
                   #IOuMouldEditor_HMI.arShotSet[#IOuMouldEditor_HMI.sSelected.sPS.iPS].Flow[#TiLoop] := #IOuMouldEditor_HMI.sSelected.sPS.arFlow[#TiLoop];
                   //Sum new Flow
                   #OUTrSumFlow := 0;

                   FOR #TiLoop_Flow := 1 TO #TiComponentAmount DO
                       #OUTrSumFlow := #OUTrSumFlow + #IOuMouldEditor_HMI.arShotSet[#IOuMouldEditor_HMI.sSelected.sPS.iPS].Flow[#TiLoop_Flow];
                   END_FOR;

                   // changed flow is not ref comp
                   IF #TiLoop <> #IOuMouldEditor_HMI.sSelected.sPS.RefComponent THEN
                       // New ratio for changed flow
                       #IOuMouldEditor_HMI.sSelected.sPS.arRatio[#TiLoop] := #IOuMouldEditor_HMI.sSelected.sPS.arFlow[#TiLoop] /
                       #IOuMouldEditor_HMI.arShotSet[#IOuMouldEditor_HMI.sSelected.sPS.iPS].Flow[#IOuMouldEditor_HMI.sSelected.sPS.RefComponent] / 100.0;
                       // changed flow is ref comp    
                   ELSE
                       // New ratio for all other flowrates
                       FOR #TiLoop_Flow := 1 TO #TiComponentAmount DO
                           IF #TiLoop_Flow <> #IOuMouldEditor_HMI.sSelected.sPS.RefComponent THEN
                               IF #IOuMouldEditor_HMI.arShotSet[#IOuMouldEditor_HMI.sSelected.sPS.iPS].Flow[#IOuMouldEditor_HMI.sSelected.sPS.RefComponent] <> 0 THEN
                                   #IOuMouldEditor_HMI.sSelected.sPS.arRatio[#TiLoop_Flow] := #IOuMouldEditor_HMI.sSelected.sPS.arFlow[#TiLoop_Flow] /
                                   #IOuMouldEditor_HMI.arShotSet[#IOuMouldEditor_HMI.sSelected.sPS.iPS].Flow[#IOuMouldEditor_HMI.sSelected.sPS.RefComponent] / 100.0;
                               ELSE
                                   #IOuMouldEditor_HMI.sSelected.sPS.arRatio[#TiLoop_Flow] := 0;
                                   #IOuMouldEditor_HMI.sSelected.sPS.arFlow[#TiLoop_Flow] := 0;
                                   #IOuMouldEditor_HMI.arShotSet[#IOuMouldEditor_HMI.sSelected.sPS.iPS].Flow[#TiLoop_Flow] := 0;
                               END_IF;
                           END_IF;
                       END_FOR;
                   END_IF;

                   //Sum new Flow
                   #OUTrSumFlow := 0;

                   FOR #TiLoop_Flow := 1 TO #TiComponentAmount DO
                       #OUTrSumFlow := #OUTrSumFlow + #IOuMouldEditor_HMI.arShotSet[#IOuMouldEditor_HMI.sSelected.sPS.iPS].Flow[#TiLoop_Flow];
                   END_FOR;
                   #IOuMouldEditor_HMI.sCalculatedValues.arTotalFlow[#IOuMouldEditor_HMI.sSelected.sPS.iPS] := #OUTrSumFlow;


                   // Calculate new ratio
                   // SumRatio
                   #OUTrSumRatio := 0;

                   FOR #TiLoop_Ratio := 1 TO #TiComponentAmount DO
                       #OUTrSumRatio := #OUTrSumRatio + #IOuMouldEditor_HMI.sSelected.sPS.arRatio[#TiLoop_Ratio];
                   END_FOR;

                   //  Calculation = 0 -> shot time fixed
                   IF #IOuMouldEditor_HMI.sSelected.iCalculation = 0 THEN
                       #IOuMouldEditor_HMI.arShotSet[#IOuMouldEditor_HMI.sSelected.sPS.iPS].PartWeight := #IOuMouldEditor_HMI.sCalculatedValues.arTotalFlow[#IOuMouldEditor_HMI.sSelected.sPS.iPS] * #IOuMouldEditor_HMI.arShotSet[#IOuMouldEditor_HMI.sSelected.sPS.iPS].FoamingTime;
                   END_IF;
                   // ----

                   //  Calculation = 2 -> weight fixed
                   IF #IOuMouldEditor_HMI.sSelected.iCalculation = 2 THEN
                       IF #IOuMouldEditor_HMI.sCalculatedValues.arTotalFlow[#IOuMouldEditor_HMI.sSelected.sPS.iPS] >= 0 THEN
                           #IOuMouldEditor_HMI.arShotSet[#IOuMouldEditor_HMI.sSelected.sPS.iPS].FoamingTime := #IOuMouldEditor_HMI.arShotSet[#IOuMouldEditor_HMI.sSelected.sPS.iPS].PartWeight / #IOuMouldEditor_HMI.sCalculatedValues.arTotalFlow[#IOuMouldEditor_HMI.sSelected.sPS.iPS];
                       END_IF;
                   END_IF;

                   //  Value changed + Save data for the last cycle to recognize changes of the values
                   #IOuMouldEditor_HMI.sStatusBits.xValueChanged := TRUE;
                   #SuMouldEditor_HMI := #IOuMouldEditor_HMI;
                   EXIT;
                   // ----

               END_IF
               ;
           END_FOR;
       END_REGION
       //_________________________________________________________________________________    
       REGION Pressure - changed
           FOR #TiLoop := 1 TO #TiComponentAmount DO
               IF #IOuMouldEditor_HMI.sSelected.sPS.arPressure[#TiLoop] <> #SuMouldEditor_HMI.sSelected.sPS.arPressure[#TiLoop] THEN

                   #IOuMouldEditor_HMI.arShotSet[#IOuMouldEditor_HMI.sSelected.sPS.iPS].Pressure[#TiLoop] := #IOuMouldEditor_HMI.sSelected.sPS.arPressure[#TiLoop];

                   //  Value changed + Save data for the last cycle to recognize changes of the values
                   #IOuMouldEditor_HMI.sStatusBits.xValueChanged := TRUE;
                   #SuMouldEditor_HMI := #IOuMouldEditor_HMI;
                   EXIT;
                   // ----

               END_IF
               ;
           END_FOR;
       END_REGION
       //_________________________________________________________________________________    
       REGION Reference component - changed
           IF #IOuMouldEditor_HMI.sSelected.sPS.RefComponent <> #SuMouldEditor_HMI.sSelected.sPS.RefComponent THEN

               #IOuMouldEditor_HMI.arShotSet[#IOuMouldEditor_HMI.sSelected.sPS.iPS].RefComponent := #IOuMouldEditor_HMI.sSelected.sPS.RefComponent;

               IF #IOuMouldEditor_HMI.sSelected.sPS.arFlow[#IOuMouldEditor_HMI.sSelected.sPS.RefComponent] = 0 THEN
                   #IOuMouldEditor_HMI.sSelected.sPS.arRatio[#IOuMouldEditor_HMI.sSelected.sPS.RefComponent] := 100.00;
               END_IF;

               // Calculation of flow in "Mixing ratio - changed"
               //  Value changed + Save data for the last cycle to recognize changes of the values
               #IOuMouldEditor_HMI.sStatusBits.xValueChanged := TRUE;
               //#SuMouldEditor_HMI := #IOuMouldEditor_HMI;

           END_IF;
       END_REGION
       //_________________________________________________________________________________    
       REGION Mixing ratio - changed
           FOR #TiLoop := 1 TO #TiComponentAmount DO
               IF #IOuMouldEditor_HMI.sSelected.sPS.arRatio[#TiLoop] <> #SuMouldEditor_HMI.sSelected.sPS.arRatio[#TiLoop] THEN

                   // only change single flow rates!
                   // SumRatio
                   #OUTrSumRatio := 0;

                   FOR #TiLoop_Ratio := 1 TO #TiComponentAmount DO
                       #OUTrSumRatio := #OUTrSumRatio + #IOuMouldEditor_HMI.sSelected.sPS.arRatio[#TiLoop_Ratio];
                   END_FOR;

                   FOR #TiLoop_Flow := 1 TO #TiComponentAmount DO

                       #IOuMouldEditor_HMI.sSelected.sPS.arFlow[#TiLoop_Flow] := #IOuMouldEditor_HMI.sCalculatedValues.arTotalFlow[#IOuMouldEditor_HMI.sSelected.sPS.iPS] /
                       #OUTrSumRatio * #IOuMouldEditor_HMI.sSelected.sPS.arRatio[#TiLoop_Flow];
                       #IOuMouldEditor_HMI.arShotSet[#IOuMouldEditor_HMI.sSelected.sPS.iPS].Flow[#TiLoop_Flow] := #IOuMouldEditor_HMI.sSelected.sPS.arFlow[#TiLoop_Flow];
                   END_FOR;

                   //  Value changed + Save data for the last cycle to recognize changes of the values
                   #IOuMouldEditor_HMI.sStatusBits.xValueChanged := TRUE;
                   #SuMouldEditor_HMI := #IOuMouldEditor_HMI;
                   EXIT;
                   // ----

               END_IF
               ;
           END_FOR;
       END_REGION
       //_________________________________________________________________________________    
       REGION Mixing head - changed
           FOR #TiLoop_PS := 1 TO #TiPartShotAmount DO
               IF #IOuMouldEditor_HMI.arShotSet[#TiLoop_PS].MHNo <> #SuMouldEditor_HMI.arShotSet[#TiLoop_PS].MHNo THEN
                   // Check if ref comp is available at this MH. Reset all values for not used components            

                   IF #RefComp > #TiComponentAmount THEN
                       #IOuMouldEditor_HMI.arShotSet[#TiLoop_PS].RefComponent := 1;
                   END_IF;

                   IF #TiComponentAmount < 6 THEN
                       FOR #TiLoop := #TiComponentAmount + 1 TO 6 DO
                           #IOuMouldEditor_HMI.arShotSet[#TiLoop_PS].Pressure[#TiLoop] := 0;
                           #IOuMouldEditor_HMI.arShotSet[#TiLoop_PS].Flow[#TiLoop] := 0;
                       END_FOR;
                   END_IF;
                   //  Value changed + Save data for the last cycle to recognize changes of the values
                   #IOuMouldEditor_HMI.sStatusBits.xValueChanged := TRUE;
                   #SuMouldEditor_HMI := #IOuMouldEditor_HMI;
                   EXIT;
                   // ----

               END_IF;
           END_FOR;
       END_REGION
       //_________________________________________________________________________________    
       REGION Two point adjust changed
           // IF #IOuMouldEditor_HMI.sSelected.sPS."2PoinMovement_Comp01" <> #SuMouldEditor_HMI.sSelected.sPS."2PoinMovement_Comp01" OR
           //     #IOuMouldEditor_HMI.sSelected.sPS."2PoinMovement_Comp02" <> #SuMouldEditor_HMI.sSelected.sPS."2PoinMovement_Comp02" OR
           //     #IOuMouldEditor_HMI.sSelected.sPS."2PoinMovement_Comp03" <> #SuMouldEditor_HMI.sSelected.sPS."2PoinMovement_Comp03" OR
           //     #IOuMouldEditor_HMI.sSelected.sPS."2PoinMovement_Comp04" <> #SuMouldEditor_HMI.sSelected.sPS."2PoinMovement_Comp04" OR
           //     #IOuMouldEditor_HMI.sSelected.sPS."2PoinMovement_Comp05" <> #SuMouldEditor_HMI.sSelected.sPS."2PoinMovement_Comp05" OR
           //     #IOuMouldEditor_HMI.sSelected.sPS."2PoinMovement_Comp06" <> #SuMouldEditor_HMI.sSelected.sPS."2PoinMovement_Comp06"
           // THEN
           //     #IOuMouldEditor_HMI.arShotSet[#IOuMouldEditor_HMI.sSelected.sPS.iPS]."2PoinMovement_Comp01" := #IOuMouldEditor_HMI.sSelected.sPS."2PoinMovement_Comp01";
           //     #IOuMouldEditor_HMI.arShotSet[#IOuMouldEditor_HMI.sSelected.sPS.iPS]."2PoinMovement_Comp02" := #IOuMouldEditor_HMI.sSelected.sPS."2PoinMovement_Comp02";
           //     #IOuMouldEditor_HMI.arShotSet[#IOuMouldEditor_HMI.sSelected.sPS.iPS]."2PoinMovement_Comp03" := #IOuMouldEditor_HMI.sSelected.sPS."2PoinMovement_Comp03";
           //     #IOuMouldEditor_HMI.arShotSet[#IOuMouldEditor_HMI.sSelected.sPS.iPS]."2PoinMovement_Comp04" := #IOuMouldEditor_HMI.sSelected.sPS."2PoinMovement_Comp04";
           //     #IOuMouldEditor_HMI.arShotSet[#IOuMouldEditor_HMI.sSelected.sPS.iPS]."2PoinMovement_Comp05" := #IOuMouldEditor_HMI.sSelected.sPS."2PoinMovement_Comp05";
           //     #IOuMouldEditor_HMI.arShotSet[#IOuMouldEditor_HMI.sSelected.sPS.iPS]."2PoinMovement_Comp06" := #IOuMouldEditor_HMI.sSelected.sPS."2PoinMovement_Comp06";

           //     //  Value changed + Save data for the last cycle to recognize changes of the values
           //     #IOuMouldEditor_HMI.sStatusBits.xValueChanged := TRUE;
           //     #SuMouldEditor_HMI := #IOuMouldEditor_HMI;
           //     // ----
           // END_IF;
       END_REGION
       //_________________________________________________________________________________    
       REGION Values in shot settings - changed
           FOR #TiLoop_PS := 1 TO #TiPartShotAmount DO
               IF #IOuMouldEditor_HMI.arShotSet[#TiLoop_PS].MHNo <> #SuMouldEditor_HMI.arShotSet[#TiLoop_PS].MHNo OR
                   #IOuMouldEditor_HMI.arShotSet[#TiLoop_PS].CP_ThrottleGap <> #SuMouldEditor_HMI.arShotSet[#TiLoop_PS].CP_ThrottleGap OR
                   #IOuMouldEditor_HMI.arShotSet[#TiLoop_PS].CP_ThrottleGap <> #SuMouldEditor_HMI.arShotSet[#TiLoop_PS].CP_ThrottleGap OR
                   #IOuMouldEditor_HMI.arShotSet[#TiLoop_PS].PartShotDisable <> #SuMouldEditor_HMI.arShotSet[#TiLoop_PS].PartShotDisable OR
                   #IOuMouldEditor_HMI.arShotSet[#TiLoop_PS].CPMoveAfterShot <> #SuMouldEditor_HMI.arShotSet[#TiLoop_PS].CPMoveAfterShot OR
                   #IOuMouldEditor_HMI.arShotSet[#TiLoop_PS].PartCounter <> #SuMouldEditor_HMI.arShotSet[#TiLoop_PS].PartCounter
               THEN

                   //  Value changed + Save data for the last cycle to recognize changes of the values
                   #IOuMouldEditor_HMI.sStatusBits.xValueChanged := TRUE;
                   #SuMouldEditor_HMI := #IOuMouldEditor_HMI;
                   EXIT;
                   // ----

               END_IF
               ;
           END_FOR;
       END_REGION
       //_________________________________________________________________________________    
       REGION Partial shot number -> copy all data
           FOR #TiLoop := 1 TO #TiComponentAmount DO
               #IOuMouldEditor_HMI.sSelected.sPS.arFlow[#TiLoop] := #IOuMouldEditor_HMI.arShotSet[#IOuMouldEditor_HMI.sSelected.sPS.iPS].Flow[#TiLoop];
               #IOuMouldEditor_HMI.sSelected.sPS.arPressure[#TiLoop] := #IOuMouldEditor_HMI.arShotSet[#IOuMouldEditor_HMI.sSelected.sPS.iPS].Pressure[#TiLoop];
           END_FOR;
       END_REGION
       //_________________________________________________________________________________    
       REGION Reference component = 100%
           #RefComp := LIMIT(MN := 1, IN := #IOuMouldEditor_HMI.sSelected.sPS.RefComponent, MX := #TiComponentAmount);
           #IOuMouldEditor_HMI.sSelected.sPS.RefComponent := #RefComp;
           #TrFlowRefComp := #IOuMouldEditor_HMI.sSelected.sPS.arFlow[#IOuMouldEditor_HMI.sSelected.sPS.RefComponent];
       END_REGION
       //_________________________________________________________________________________    
       REGION Calculate ration out OF flow rate
           FOR #TiLoop := 1 TO #TiComponentAmount DO
               IF #TiLoop = #IOuMouldEditor_HMI.sSelected.sPS.RefComponent THEN
                   #IOuMouldEditor_HMI.sSelected.sPS.arRatio[#TiLoop] := 100.00;
               ELSE
                   IF #TrFlowRefComp > 00 THEN
                       #IOuMouldEditor_HMI.sSelected.sPS.arRatio[#TiLoop] := #IOuMouldEditor_HMI.sSelected.sPS.arFlow[#TiLoop] /
                       #TrFlowRefComp * 100.0;
                   END_IF;
               END_IF;
           END_FOR;
       END_REGION
       //_________________________________________________________________________________    
       #IOuMouldEditor_HMI.sSelected.sPS.RefComponent := #IOuMouldEditor_HMI.arShotSet[#IOuMouldEditor_HMI.sSelected.sPS.iPS].RefComponent;
       //_________________________________________________________________________________    
       REGION Safe changes
           // Check min/max shot time and max flowrates for each component. If out of range ask for change or discard changes   
           IF #IOuMouldEditor_HMI.sStatusBits.xSafeChanges THEN
               FOR #TiLoop_PS := 1 TO #TiPartShotAmount DO
                   // check total flow or total weight is zero
                   IF #IOuMouldEditor_HMI.sCalculatedValues.arTotalFlow[#TiLoop_PS] = 0 OR #IOuMouldEditor_HMI.arShotSet[#TiLoop_PS].PartWeight = 0 THEN
                       #IOuMouldEditor_HMI.sStatusBits.xFaultValuesnotvalid := TRUE;
                   END_IF;
                   // check foaming time for all partshots
                   IF #IOuMouldEditor_HMI.arShotSet[#TiLoop_PS].FoamingTime < "InterfaceVisu".MinShottime OR #IOuMouldEditor_HMI.arShotSet[#TiLoop_PS].FoamingTime > "InterfaceVisu".MaxShottime THEN
                       #IOuMouldEditor_HMI.sStatusBits.xFaultValuesnotvalid := TRUE;
                   END_IF;
                   // check flow rate for all part shots
                   FOR #TiLoop_Flow := 1 TO #TiComponentAmount DO
                       // Maximum flow rate limit reached
                       IF #IOuMouldEditor_HMI.arShotSet[#TiLoop_PS].Flow[#TiLoop_Flow] > "InterfaceVisu".MaxFlow[#TiLoop_Flow] THEN
                           #IOuMouldEditor_HMI.sStatusBits.xFaultValuesnotvalid := TRUE;
                       END_IF;
                       // Minimum flow rate limit reached
                       IF #IOuMouldEditor_HMI.arShotSet[#TiLoop_PS].Flow[#TiLoop_Flow] < "InterfaceVisu".MinFlow[#TiLoop_Flow] AND
                           #IOuMouldEditor_HMI.arShotSet[#TiLoop_PS].Flow[#TiLoop_Flow] <> 0 THEN
                           #IOuMouldEditor_HMI.sStatusBits.xFaultValuesnotvalid := TRUE;
                       END_IF;

                   END_FOR;

               END_FOR;
               #IOuMouldEditor_HMI.sStatusBits.xSafeChanges := FALSE;

               IF #IOuMouldEditor_HMI.sStatusBits.xFaultValuesnotvalid = FALSE THEN
                   #IOuMouldEditor_HMI.sStatusBits.xValueChanged := FALSE;
                   #IOuMouldEditor_HMI.sStatusBits.xSafeChanges := FALSE;
                   #IOuMouldEditor_HMI.sStatusBits.xDiscardChanges := FALSE;

                   FOR #TiLoop_PS := 1 TO #TiPartShotAmount DO
                       // When the selected Tool less or equal 100 is, transfer the values to DB925
                       IF #IOuMouldEditor_HMI.sSelected.iTool <= "AmountToolsDB" THEN
                           "DB925_ShotData_1".Tool[#IOuMouldEditor_HMI.sSelected.iTool].Shot[#TiLoop_PS] := #IOuMouldEditor_HMI.arShotSet[#TiLoop_PS];
                       END_IF;
                       // When the selected Tool bigger than 100 and less or equal 200 is, transfer the values to DB926
                       IF #IOuMouldEditor_HMI.sSelected.iTool > "AmountToolsDB" AND #IOuMouldEditor_HMI.sSelected.iTool <= (2*"AmountToolsDB") THEN
                           "DB926_ShotData_2".Tool[#IOuMouldEditor_HMI.sSelected.iTool-"AmountToolsDB"].Shot[#TiLoop_PS] := #IOuMouldEditor_HMI.arShotSet[#TiLoop_PS];
                       END_IF;
                   END_FOR;

                   "DB930_Tools".Tool[#IOuMouldEditor_HMI.sSelected.iTool] := #IOuMouldEditor_HMI.uTools;
               END_IF;
           END_IF;
       END_REGION
       //_________________________________________________________________________________    
       REGION Delete program
           IF #IOuMouldEditor_HMI.sStatusBits.xDeleteProgram THEN
               #IOuMouldEditor_HMI.sStatusBits.xDeleteProgram := false;
               "FC4_Check_allocation"(Selected_tool:=#IOuMouldEditor_HMI.sSelected.iTool,
                                      Delete_not_allowed=>#IOuMouldEditor_HMI.sStatusBits.xFaultDeleteProgram);

               IF NOT #IOuMouldEditor_HMI.sStatusBits.xFaultDeleteProgram THEN
                   #IOuMouldEditor_HMI.uTools.PartShot_Amount := 0;
                   #Nullbyte := 0;
                   // Delete tool data
                   // When the selected Tool less or equal 100 is, transfer the values to DB925
                   IF #IOuMouldEditor_HMI.sSelected.iTool <= "AmountToolsDB" THEN
                       #Retval := FILL(BVAL := #Nullbyte, BLK => "DB925_ShotData_1".Tool[#IOuMouldEditor_HMI.sSelected.iTool]);
                   END_IF;
                   // When the selected Tool bigger than 100 and less or equal 200 is, transfer the values to DB926
                   IF #IOuMouldEditor_HMI.sSelected.iTool > "AmountToolsDB" AND #IOuMouldEditor_HMI.sSelected.iTool <= (2 * "AmountToolsDB") THEN
                       #Retval := FILL(BVAL := #Nullbyte, BLK => "DB926_ShotData_2".Tool[#IOuMouldEditor_HMI.sSelected.iTool-"AmountToolsDB"]);
                   END_IF;

                   #Retval := FILL(BVAL := #Nullbyte, BLK => "DB930_Tools".Tool[#IOuMouldEditor_HMI.sSelected.iTool]);
                   #Retval := FILL(BVAL := #Nullbyte, BLK => #IOuMouldEditor_HMI.arShotSet);
                   "DB930_Tools".Tool[#IOuMouldEditor_HMI.sSelected.iTool].tool_name := '';
               END_IF;

           END_IF;
       END_REGION
       //_________________________________________________________________________________    
       REGION Save data FOR the last cycle TO recognize changes OF the values
           #SuMouldEditor_HMI := #IOuMouldEditor_HMI;
       END_REGION
       //_________________________________________________________________________________    
       REGION Visibility OF part shots AND "grey" fields FOR NOT changing settings
           // Column
           // Column - shot time blocked
           IF #IOuMouldEditor_HMI.sSelected.iCalculation = 0 THEN   // Statement section REGION
               #IOuMouldEditor_HMI.sColumn.iShotTime := #IOuMouldEditor_HMI.uTools.PartShot_Amount;
           ELSE
               #IOuMouldEditor_HMI.sColumn.iShotTime := 0;
           END_IF;

           // Column - total flow blocked
           IF #IOuMouldEditor_HMI.sSelected.iCalculation = 1 THEN   // Statement section REGION
               #IOuMouldEditor_HMI.sColumn.iTotalFlow := #IOuMouldEditor_HMI.uTools.PartShot_Amount;
           ELSE
               #IOuMouldEditor_HMI.sColumn.iTotalFlow := 0;
           END_IF;

           // Column - total weight blocked
           IF #IOuMouldEditor_HMI.sSelected.iCalculation = 2 THEN   // Statement section REGION
               #IOuMouldEditor_HMI.sColumn.iTotalWeight := #IOuMouldEditor_HMI.uTools.PartShot_Amount;
           ELSE
               #IOuMouldEditor_HMI.sColumn.iTotalWeight := 0;
           END_IF;

           // Row - Visibility of change partial shot
           FOR #TiLoop := 1 TO "AmountPartShots" DO
               IF #TiLoop <> #IOuMouldEditor_HMI.sSelected.sPS.iPS AND
                   #TiLoop <= BYTE_TO_INT(#IOuMouldEditor_HMI.uTools.PartShot_Amount)
               THEN
                   #IOuMouldEditor_HMI.sRow.arChangePartialShot[#TiLoop] := TRUE;
               ELSE
                   #IOuMouldEditor_HMI.sRow.arChangePartialShot[#TiLoop] := FALSE;
               END_IF;

           END_FOR;
       END_REGION
   END_IF;
END_FUNCTION_BLOCK

FUNCTION_BLOCK "FB009_Faults"   // FB9, STL
TITLE = Faults indication of machines and plant
{ S7_Optimized_Access := 'FALSE' }
AUTHOR : KT242
VERSION : 0.1
   VAR_TEMP
      Stoe_Quitt : Bool;
      Quitt : Bool;
   END_VAR
BEGIN

REGION Network 1
   //      O     "E0.4QuitFault"
   //      O     "Tag_7"
   //      =     "E0.4QuitFault"
END_REGION

REGION Network 2: Bits of fault levels
         A     "DB009_Faults".Faults_FKT_Grp_1_M1;
         =     "DB009_Faults".Fault_State_Grp_1_M1;
         A     "DB009_Faults".Faults_FKT_Grp_2_M1;
         =     "DB009_Faults".Fault_State_Grp_2_M1;
         A     "DB009_Faults".Faults_FKT_Grp_3_M1;
         =     "DB009_Faults".Fault_State_Grp_3_M1;

         A     "DB009_Faults".Faults_FKT_Grp_1_M2;
         =     "DB009_Faults".Fault_State_Grp_1_M2;
         A     "DB009_Faults".Faults_FKT_Grp_2_M2;
         =     "DB009_Faults".Fault_State_Grp_2_M2;
         A     "DB009_Faults".Faults_FKT_Grp_3_M2;
         =     "DB009_Faults".Fault_State_Grp_3_M2;

         CLR;
         =     "DB009_Faults".Fault_State_Grp_1_M3;
         =     "DB009_Faults".Fault_State_Grp_2_M3;
         =     "DB009_Faults".Fault_State_Grp_3_M3;
         =     "DB009_Faults".Fault_State_Grp_1_M4;
         =     "DB009_Faults".Fault_State_Grp_2_M4;
         =     "DB009_Faults".Fault_State_Grp_3_M4;

         A     "DB009_Faults".Faults_FKT_Grp_1_ExtP;
         =     "DB009_Faults".Fault_State_Grp_1_ExtP;
         A     "DB009_Faults".Faults_FKT_Grp_2_ExtP;
         =     "DB009_Faults".Fault_State_Grp_2_ExtP;
         A     "DB009_Faults".Faults_FKT_Grp_3_ExtP;
         =     "DB009_Faults".Fault_State_Grp_2_ExtP;

         O     "T_QuitFault";
         O     "FRA_KM_Quitt";
         =     #Quitt;

         CALL  "FC089_quit_Faults"
         ( IN_Button_Acknowledge    := #Quitt,  //"T_QuitFault"
           IN_Button_Horn_Off       := FALSE,  // "E0.4QuitFault"
           IN_First_PLC_cycle       := "Flag_Erster_SPS_Zyklus",
           IN_IndicatorLampTest     := "DB619_State_MPart".Operationmode[1].Lamptest,
           IN_Fault_Grp_1_active_M1 := "DB009_Faults".Fault_State_Grp_1_M1,
           IN_Fault_Grp_2_active_M1 := "DB009_Faults".Fault_State_Grp_2_M1,
           IN_Fault_Grp_3_active_M1 := "DB009_Faults".Fault_State_Grp_3_M1,
           IN_Fault_Grp_1_active_M2 := "DB009_Faults".Fault_State_Grp_1_M2,
           IN_Fault_Grp_2_active_M2 := "DB009_Faults".Fault_State_Grp_2_M2,
           IN_Fault_Grp_3_active_M2 := "DB009_Faults".Fault_State_Grp_3_M2,
           IN_Fault_Grp_1_active_M3 := "DB009_Faults".Fault_State_Grp_1_M3,
           IN_Fault_Grp_2_active_M3 := "DB009_Faults".Fault_State_Grp_2_M3,
           IN_Fault_Grp_3_active_M3 := "DB009_Faults".Fault_State_Grp_3_M3,
           IN_Fault_Grp_1_active_M4 := "DB009_Faults".Fault_State_Grp_1_M4,
           IN_Fault_Grp_2_active_M4 := "DB009_Faults".Fault_State_Grp_2_M4,
           IN_Fault_Grp_3_active_M4 := "DB009_Faults".Fault_State_Grp_3_M4,
           IN_Fault_Grp_1_active_AP := "DB009_Faults".Fault_State_Grp_1_ExtP,
           IN_Fault_Grp_2_active_AP := "DB009_Faults".Fault_State_Grp_2_ExtP,
           IN_Fault_Grp_3_active_AP := "DB009_Faults".Fault_State_Grp_3_ExtP,
           OUT_acoustical_indicator := "H_Fault_horn_M1",
           OUT_optical_indicator    := "H_Fault_lamp_M1",
           IO_Fault_changed_M1      := "DB009_Faults".Faultschanging_M1,
           IO_Fault_changed_M2      := "DB009_Faults".Faultschanging_M2,
           IO_Fault_changed_M3      := "DB009_Faults".Faultschanging_M3,
           IO_Fault_changed_M4      := "DB009_Faults".Faultschanging_M4,
           IO_Fault_changed_AP      := "DB009_Faults".Faultschanging_ExtP,
           IO_Horn                  := "DB009_Faults".HF_Horn,
           IO_Reset_fault_Grp       := "DB009_Faults".Faults_Reset_Group,
           IO_Reset_fault_Fkt       := "DB009_Faults".Faults_Reset_FKT_M1,
           IO_Quit_Edge             := "DB009_Faults".HF_Faults_Quit
         );
   //-----
         O     "DB009_Faults".Fault_State_Grp_1_M1;
         O     "DB009_Faults".Fault_State_Grp_2_M1;
         O     "DB009_Faults".Fault_State_Grp_3_M1;
         O     "DB009_Faults".Fault_State_Grp_1_M2;
         O     "DB009_Faults".Fault_State_Grp_2_M2;
         O     "DB009_Faults".Fault_State_Grp_3_M2;
         O     "DB009_Faults".Fault_State_Grp_1_M3;
         O     "DB009_Faults".Fault_State_Grp_2_M3;
         O     "DB009_Faults".Fault_State_Grp_3_M3;
         O     "DB009_Faults".Fault_State_Grp_1_M4;
         O     "DB009_Faults".Fault_State_Grp_2_M4;
         O     "DB009_Faults".Fault_State_Grp_3_M4;
         O     "DB009_Faults".Fault_State_Grp_1_ExtP;
         O     "DB009_Faults".Fault_State_Grp_2_ExtP;
         O     "DB009_Faults".Fault_State_Grp_2_ExtP;
         =     "DB009_Faults".Fault_State_Grp_1_3_Exist;
   //-----
         A     "DB009_Faults".Faults_Reset_FKT_M1;
         S     "DB009_Faults".HF_FaultsQuitOB35;
   //-----
         A     "DB009_Faults".Faults_Reset_Group;
         R     "DB009_Faults".Faults_FKT_Grp_1_M1;
         R     "DB009_Faults".Faults_FKT_Grp_2_M1;
         R     "DB009_Faults".Faults_FKT_Grp_3_M1;
         R     "DB009_Faults".Faults_FKT_Grp_1_M2;
         R     "DB009_Faults".Faults_FKT_Grp_2_M2;
         R     "DB009_Faults".Faults_FKT_Grp_3_M2;
         R     "DB009_Faults".Faults_FKT_Grp_1_M3;
         R     "DB009_Faults".Faults_FKT_Grp_2_M3;
         R     "DB009_Faults".Faults_FKT_Grp_3_M3;
         R     "DB009_Faults".Faults_FKT_Grp_1_M4;
         R     "DB009_Faults".Faults_FKT_Grp_2_M4;
         R     "DB009_Faults".Faults_FKT_Grp_3_M4;
         R     "DB009_Faults".Faults_FKT_Grp_1_ExtP;
         R     "DB009_Faults".Faults_FKT_Grp_2_ExtP;
         R     "DB009_Faults".Faults_FKT_Grp_3_ExtP;
   //-----
END_REGION

REGION Network 3: General faults of machines
         CALL  "FC081_FaultsGen"
         ( IN_Erster_SPS_Zyklus := "Flag_Erster_SPS_Zyklus"
         );
END_REGION

REGION Network 4: Faults Profibus
         CALL  "FC082_FaultProfiBus";
END_REGION

REGION Network 5: Lamp machine ok for foaming
         O     "H_Ready_for_Operation_M1";
         O     "H_Ready_for_Operation_M2";
         =     "H_Ready_for_Operation";
END_REGION

REGION Network 6: Signalshow fault massages and messages at visu
         O     "DB009_Faults".NewMessage_M1;
         O     "DB009_Faults".GoneMessage_M1;
         O     "DB009_Faults".Faultschanging_M1;
         O     "DB009_Faults".Faults_Reset_FKT_M1;
         AN    "DB009_Faults".MessageChangedToVisu;
         S     "DB009_Faults".MessageChangedToVisu;
         R     "DB009_Faults".NewMessage_M1;
         R     "DB009_Faults".GoneMessage_M1;
         R     "DB009_Faults".MessageChangedNext;

         O     "DB009_Faults".NewMessage_M1;
         O     "DB009_Faults".GoneMessage_M1;
         O     "DB009_Faults".Faultschanging_M1;
         O     "DB009_Faults".Faults_Reset_FKT_M1;
         A     "DB009_Faults".MessageChangedToVisu;
         S     "DB009_Faults".MessageChangedNext;
END_REGION
END_FUNCTION_BLOCK

FUNCTION_BLOCK "FB011_OP_CirceMode_M1"   // FB11, STL
TITLE = Operation mode and cycle mode of machine 01
{ S7_Optimized_Access := 'FALSE' }
AUTHOR : KT242
VERSION : 0.1
   VAR_TEMP
      Temp_Release_HP : Bool;
      Temp_ShotPreperation : Bool;
      Temp_Automatic_MH1 : Bool;
      Temp_HPCirc_aft_shot_MH1 : Bool;
      Temp_HF_LP_circ : Bool;
      Temp_TestMode : Bool;
      Temp_TestA : Bool;
      Temp_TestB : Bool;
      Temp_H_TestA : Bool;
      Temp_H_TestB : Bool;
      Dummy : Bool;
   END_VAR
BEGIN

REGION Network 1: State switch service/ operation
         L     0;
         T     "DB614_MH_State".MH_Status[1].State_Service;
         T     "DB614_MH_State".MH_Status[2].State_Service;
         T     "DB614_MH_State".MH_Status[3].State_Service;
         T     "DB614_MH_State".MH_Status[4].State_Service;
         T     "DB614_MH_State".MH_Status[5].State_Service;
         T     "DB614_MH_State".MH_Status[6].State_Service;
         T     "DB614_MH_State".MH_Status[7].State_Service;
         T     "DB614_MH_State".MH_Status[8].State_Service;
         T     "DB614_MH_State".MH_Status[8].State_Service;
         T     "DB614_MH_State".MH_Status[9].State_Service;
         T     "DB614_MH_State".MH_Status[10].State_Service;
         T     "DB614_MH_State".MH_Status[11].State_Service;
         T     "DB614_MH_State".MH_Status[12].State_Service;
   //-----
         A     "DB614_MH_State".MH_Status[1].Switch_Service_ON_OFF;
         JCN   NoServ_MH01;
         L     1;
         T     "DB614_MH_State".MH_Status[1].State_Service;
   NoServ_MH01:NOP   0;
   //-----
         A     "DB614_MH_State".MH_Status[2].Switch_Service_ON_OFF;
         JCN   NoServ_MH02;
         L     1;
         T     "DB614_MH_State".MH_Status[2].State_Service;
   NoServ_MH02:NOP   0;
   //-----
         A     "DB614_MH_State".MH_Status[3].Switch_Service_ON_OFF;
         JCN   NoServ_MH03;
         L     1;
         T     "DB614_MH_State".MH_Status[3].State_Service;
   NoServ_MH03:NOP   0;
   //-----
         A     "DB614_MH_State".MH_Status[4].Switch_Service_ON_OFF;
         JCN   NoServ_MH04;
         L     1;
         T     "DB614_MH_State".MH_Status[4].State_Service;
   NoServ_MH04:NOP   0;
   //-----
         A     "DB614_MH_State".MH_Status[5].Switch_Service_ON_OFF;
         JCN   NoServ_MH05;
         L     1;
         T     "DB614_MH_State".MH_Status[5].State_Service;
   NoServ_MH05:NOP   0;
   //-----
         A     "DB614_MH_State".MH_Status[6].Switch_Service_ON_OFF;
         JCN   NoServ_MH06;
         L     1;
         T     "DB614_MH_State".MH_Status[6].State_Service;
   NoServ_MH06:NOP   0;
   //-----
         A     "DB614_MH_State".MH_Status[7].Switch_Service_ON_OFF;
         JCN   NoServ_MH07;
         L     1;
         T     "DB614_MH_State".MH_Status[7].State_Service;
   NoServ_MH07:NOP   0;
   //-----
         A     "DB614_MH_State".MH_Status[8].Switch_Service_ON_OFF;
         JCN   NoServ_MH08;
         L     1;
         T     "DB614_MH_State".MH_Status[8].State_Service;
   NoServ_MH08:NOP   0;
   //-----
         A     "DB614_MH_State".MH_Status[9].Switch_Service_ON_OFF;
         JCN   NoServ_MH09;
         L     1;
         T     "DB614_MH_State".MH_Status[9].State_Service;
   NoServ_MH09:NOP   0;
   //-----
         A     "DB614_MH_State".MH_Status[10].Switch_Service_ON_OFF;
         JCN   NoServ_MH10;
         L     1;
         T     "DB614_MH_State".MH_Status[10].State_Service;
   NoServ_MH10:NOP   0;
   //-----
         A     "DB614_MH_State".MH_Status[11].Switch_Service_ON_OFF;
         JCN   NoServ_MH11;
         L     1;
         T     "DB614_MH_State".MH_Status[11].State_Service;
   NoServ_MH11:NOP   0;
   //-----
         A     "DB614_MH_State".MH_Status[12].Switch_Service_ON_OFF;
         JCN   NoServ_MH12;
         L     1;
         T     "DB614_MH_State".MH_Status[12].State_Service;
   NoServ_MH12:NOP   0;
   //-----
END_REGION

REGION Network 2: Switch operation mode ->ON -> with foam to open mixinghead (extarnel)

         A     "DB619_State_MPart".SWU[1].Open_SWU."01";
         A     "DB614_MH_State".MH_Status[1].Switch_Service_ON_OFF;
         O;
         A     "DB619_State_MPart".SWU[1].Open_SWU."02";
         A     "DB614_MH_State".MH_Status[2].Switch_Service_ON_OFF;
         O;
         A     "DB619_State_MPart".SWU[1].Open_SWU."03";
         A     "DB614_MH_State".MH_Status[3].Switch_Service_ON_OFF;
         O;
         A     "DB619_State_MPart".SWU[1].Open_SWU."04";
         A     "DB614_MH_State".MH_Status[4].Switch_Service_ON_OFF;
         O;
         A     "DB619_State_MPart".SWU[1].Open_SWU."05";
         A     "DB614_MH_State".MH_Status[5].Switch_Service_ON_OFF;
         O;
         A     "DB619_State_MPart".SWU[1].Open_SWU."06";
         A     "DB614_MH_State".MH_Status[6].Switch_Service_ON_OFF;
         O;
         A     "DB619_State_MPart".SWU[1].Open_SWU."07";
         A     "DB614_MH_State".MH_Status[7].Switch_Service_ON_OFF;
         O;
         A     "DB619_State_MPart".SWU[1].Open_SWU."08";
         A     "DB614_MH_State".MH_Status[8].Switch_Service_ON_OFF;
         O;
         A     "DB619_State_MPart".SWU[1].Open_SWU."09";
         A     "DB614_MH_State".MH_Status[9].Switch_Service_ON_OFF;
         O;
         A     "DB619_State_MPart".SWU[1].Open_SWU."10";
         A     "DB614_MH_State".MH_Status[10].Switch_Service_ON_OFF;
         O;
         A     "DB619_State_MPart".SWU[1].Open_SWU."11";
         A     "DB614_MH_State".MH_Status[11].Switch_Service_ON_OFF;
         O;
         A     "DB619_State_MPart".SWU[1].Open_SWU."12";
         A     "DB614_MH_State".MH_Status[12].Switch_Service_ON_OFF;
         =     "DB619_State_MPart".Operationmode[1].SwitchOperation;
END_REGION

REGION Network 3: Test shot Sonder
         L     0;
         T     "DB614_MH_State".MH_Status[1].State_Testshot_A;
         T     "DB614_MH_State".MH_Status[1].State_Testshot_B;

         AN    "DB123_MH_IO_Signals".MH[1].IN.MH_Manual_Mode;
         R     "DB614_MH_State".MH_Status[1].Switch_Testshot_A_ON_OFF;
         R     "DB614_MH_State".MH_Status[1].Switch_Testshot_B_ON_OFF;

         A     "DB614_MH_State".MH_Status[1].Switch_Testshot_A_ON_OFF;
         JCN   TestA_MH01;
         L     1;
         T     "DB614_MH_State".MH_Status[1].State_Testshot_A;
         L     0;
         T     "DB614_MH_State".MH_Status[1].State_Testshot_B;
   TestA_MH01:NOP   0;

         A     "DB614_MH_State".MH_Status[1].Switch_Testshot_B_ON_OFF;
         JCN   TestB_MH01;
         L     1;
         T     "DB614_MH_State".MH_Status[1].State_Testshot_B;
         L     0;
         T     "DB614_MH_State".MH_Status[1].State_Testshot_A;
   TestB_MH01:NOP   0;

         A     "DB614_MH_State".MH_Status[1].Switch_Testshot_A_ON_OFF;
         O     "DB614_MH_State".MH_Status[1].Switch_Testshot_B_ON_OFF;
         =     #Temp_TestMode;

         A     "DB614_MH_State".MH_Status[1].Switch_Testshot_A_ON_OFF;
         A     "DB123_MH_IO_Signals".MH[1].IN.MH_Start;
         =     #Temp_TestA;

         A     "DB614_MH_State".MH_Status[1].Switch_Testshot_B_ON_OFF;
         A     "DB123_MH_IO_Signals".MH[1].IN.MH_Start;
         =     #Temp_TestB;

         A     "DB009_Faults".Faults_FKT_Grp_1_M1;
         L     s5t#3s;
         SP    "TM_Group1_Fault";

         A     #Temp_TestMode;
         A     "DB619_State_MPart".Cycle[1].running;
         AN    "DB614_MH_State".MH_Status[1].Switch_Testshot_A_ON_OFF;
         O     "DB123_MH_IO_Signals".MH[1].OUT.MH.V_LowPressure_Circ_MH;
         O     "TM_Group1_Fault";
   //      NOT
         =     "V_Bypass_C1";

         A     #Temp_TestMode;
         A     "DB619_State_MPart".Cycle[1].running;
         AN    "DB614_MH_State".MH_Status[1].Switch_Testshot_B_ON_OFF;
         O     "DB123_MH_IO_Signals".MH[1].OUT.MH.V_LowPressure_Circ_MH;
         O     "TM_Group1_Fault";
   //      NOT
         =     "V_Bypass_C2";
END_REGION

REGION Network 4: Auslitern
         CALL  "FC115_Testen"
         ( IN_Betriebsart_Testen   := "DB619_State_MPart".Operationmode[1].Test,
           IN_Betriebsart_Betrieb  := "DB619_State_MPart".Operationmode[1].Operation,
           IN_Lampentest           := FALSE,
           IN_Start_Testen_K1      := #Temp_TestA,
           IN_Start_Testen_K2      := #Temp_TestB,
           IN_Start_Testen_K3      := FALSE,
           IN_Start_Testen_K4      := FALSE,
           IN_Stop_Testen          := "DB123_MH_IO_Signals".MH[1].IN.MH_Stop,
           IN_Stoerung_Gruppe_1    := "DB009_Faults".Faults_FKT_Grp_1_M1,
           IN_Zyklus_Freigabe      := "DB619_State_MPart".Cycle[1].Release,
           IN_Zyklus_laeuft        := "DB619_State_MPart".ToolMa[1].StationActive,
           IN_Zyklus_Schuss_laeuft := "DB619_State_MPart".Cycle[1].ShotRuns,
           IN_Imp_Zyklus_Ende      := "DB619_State_MPart".Cycle[1].Pulse_ToolFinished,
           IN_Zyklus_KLZ2_u_ff     := "DB619_State_MPart".Cycle[1].LastStanbyTimeTool,
           OUT_H_Testen_K1         := #Temp_H_TestA,
           OUT_H_Testen_K2         := #Temp_H_TestB,
           OUT_H_Testen_K3         := #Dummy,
           OUT_H_Testen_K4         := #Dummy,
           OUT_V_Testen_K1         := #Dummy,
           OUT_V_Testen_K2         := #Dummy,
           OUT_V_Testen_K3         := #Dummy,
           OUT_V_Testen_K4         := #Dummy,
           IO_Status               := "DB110_Interf_Program_M1".Test_M01
         );
   //
         A     "DB110_Interf_Program_M1".Test_M01.Test_K2;
         =     "Duese_K1_MH01";

         A     "DB110_Interf_Program_M1".Test_M01.Test_K1;
         =     "Duese_K2_MH01";

         A     #Temp_H_TestA;
         O     #Temp_H_TestB;
         =     "DB110_Interf_Program_M1".Test_M01.Spare_0_7;
END_REGION

REGION Network 5: Detecting operation modes
   //-----
         CALL  "FC011_OperationMode"
         ( IN_ContrVoltage        := "Controlvoltage",
           IN_Connection_OK       := TRUE,
           IN_SS_Manual           := "S_OM_Manual",
           IN_SS_Auto             := "S_OM_Auto",
           IN_SS_Test             := #Temp_TestMode,  //"S_OM_Test"
           IN_LampTest            := FALSE,  // "T_Lampentest"
           IN_Cycle_selected      := "DB619_State_MPart".Recirculation[1].Is_selected,
           IN_SS_CylinderService  := "DB619_State_MPart".CylinderManager[1].Cylinderservice,
           IN_Hydraulic_OK        := "DB619_State_MPart".Machine[1].HydStartUp_finished,
           IN_OperationMode_Timer := "TM_OM_M1",
           IO_Status              := "DB619_State_MPart".Operationmode[1]
         );
   //-----
END_REGION

REGION Network 6: High pressure cycle after automatic shot
   //-----
         A     "DB123_MH_IO_Signals".MH[1].IN.MH_Auto_Mode;
         A     "DB619_State_MPart".SWU[1].Open_SWU_allone."01";
   //     CLR
         =     #Temp_Automatic_MH1;
   //-----
         A     "DB619_State_MPart".Cycle[1].ShotRuns;
         A     #Temp_Automatic_MH1;
         L     "DB700_Machine".Machine[1].HP_time_after_shot;
         SF    "TM_HP_after_shot_M1";
   //-----
         O     "TM_HP_after_shot_M1";
   //      CLR
         =     "DB619_State_MPart".Machine[1].HP_after_shot;
   //-----
         A(;
         O     "DB619_State_MPart".Machine[1].HP_after_shot;
         FP    "DB619_State_MPart".Machine[1].Flag_P_HP_after_shot;
         );
         AN    "DB619_State_MPart".Recirculation[1].HP_is_active;
         O;
         A(;
         A     "DB619_State_MPart".Machine[1].HP_after_shot;
         FN    "DB619_State_MPart".Machine[1].Flag_N_HP_after_shot;
         );
         A     "DB619_State_MPart".Recirculation[1].HP_is_active;
         =     #Temp_HPCirc_aft_shot_MH1;
   //-----
         A     #Temp_Automatic_MH1;
         JC    M001;
         L     S5T#0MS;
         CLR;
         SP    "TM_HP_after_shot_M1";
   M001: NOP   0;
   //-----
END_REGION

REGION Network 7: Release of high pressure cycle
         O     "DB619_State_MPart".Machine[1].HP_after_shot;
         ON    "DB619_State_MPart".Cycle[1].running;
         A     "DB619_State_MPart".Operationmode[1].Active;
         AN    "DB009_Faults".Fault_State_Grp_1_M1;
         =     #Temp_Release_HP;
   //-----
END_REGION

REGION Network 8: Select high pressure cycle by PUC08 or mixinghead panel
   //__________________________________________________________________
   // Select high pressure mixinghead 01:
   // ------------------------------------
         O     #Temp_HPCirc_aft_shot_MH1;
         O     "DB123_MH_IO_Signals".MH[1].IN.MH_HP_Circ_MH;
         O     "DB614_MH_State".MH_Status[1].Switch_HP_ON_OFF;
         =     "DB619_State_MPart".Recirculation[1].Button_HP."01";
   //__________________________________________________________________
   //Select high pressure mixinghead 02:
   //------------------------------------
         O     "DB123_MH_IO_Signals".MH[2].IN.MH_HP_Circ_MH;
         O     "DB614_MH_State".MH_Status[2].Switch_HP_ON_OFF;
         =     "DB619_State_MPart".Recirculation[1].Button_HP."02";
   //__________________________________________________________________
   //Select high pressure mixinghead 03:
   //------------------------------------
         O     "DB123_MH_IO_Signals".MH[3].IN.MH_HP_Circ_MH;
         O     "DB614_MH_State".MH_Status[3].Switch_HP_ON_OFF;
         =     "DB619_State_MPart".Recirculation[1].Button_HP."03";
   //__________________________________________________________________
   //Select high pressure mixinghead 04:
   //------------------------------------
         O     "DB123_MH_IO_Signals".MH[4].IN.MH_HP_Circ_MH;
         O     "DB614_MH_State".MH_Status[4].Switch_HP_ON_OFF;
         =     "DB619_State_MPart".Recirculation[1].Button_HP."04";
   //__________________________________________________________________
   //Select high pressure mixinghead 05:
   //------------------------------------
         O     "DB123_MH_IO_Signals".MH[5].IN.MH_HP_Circ_MH;
         O     "DB614_MH_State".MH_Status[5].Switch_HP_ON_OFF;
         =     "DB619_State_MPart".Recirculation[1].Button_HP."05";
   //__________________________________________________________________
   //Select high pressure mixinghead 06:
   //------------------------------------
         O     "DB123_MH_IO_Signals".MH[6].IN.MH_HP_Circ_MH;
         O     "DB614_MH_State".MH_Status[6].Switch_HP_ON_OFF;
         =     "DB619_State_MPart".Recirculation[1].Button_HP."06";
   //__________________________________________________________________
   //Select high pressure mixinghead 07:
   //------------------------------------
         O     "DB123_MH_IO_Signals".MH[7].IN.MH_HP_Circ_MH;
         O     "DB614_MH_State".MH_Status[7].Switch_HP_ON_OFF;
         =     "DB619_State_MPart".Recirculation[1].Button_HP."07";
   //__________________________________________________________________
   //Select high pressure mixinghead 08:
   //------------------------------------
         O     "DB123_MH_IO_Signals".MH[8].IN.MH_HP_Circ_MH;
         O     "DB614_MH_State".MH_Status[8].Switch_HP_ON_OFF;
         =     "DB619_State_MPart".Recirculation[1].Button_HP."08";
   //__________________________________________________________________
   //Select high pressure mixinghead 09:
   //------------------------------------
         O     "DB123_MH_IO_Signals".MH[9].IN.MH_HP_Circ_MH;
         O     "DB614_MH_State".MH_Status[9].Switch_HP_ON_OFF;
         =     "DB619_State_MPart".Recirculation[1].Button_HP."09";
   //__________________________________________________________________
   //Select high pressure mixinghead 10:
   //------------------------------------
         O     "DB123_MH_IO_Signals".MH[10].IN.MH_HP_Circ_MH;
         O     "DB614_MH_State".MH_Status[10].Switch_HP_ON_OFF;
         =     "DB619_State_MPart".Recirculation[1].Button_HP."10";
   //__________________________________________________________________
   //Select high pressure mixinghead 11:
   //------------------------------------
         O     "DB123_MH_IO_Signals".MH[11].IN.MH_HP_Circ_MH;
         O     "DB614_MH_State".MH_Status[11].Switch_HP_ON_OFF;
         =     "DB619_State_MPart".Recirculation[1].Button_HP."11";
   //__________________________________________________________________
   //Select high pressure mixinghead 12:
   //------------------------------------
         O     "DB123_MH_IO_Signals".MH[12].IN.MH_HP_Circ_MH;
         O     "DB614_MH_State".MH_Status[12].Switch_HP_ON_OFF;
         =     "DB619_State_MPart".Recirculation[1].Button_HP."12";
   //__________________________________________________________________
   //
END_REGION

REGION Network 9: Reset the HP switches at the Panel
         SET;
         R     "DB614_MH_State".MH_Status[0].Switch_HP_ON_OFF;
         R     "DB614_MH_State".MH_Status[1].Switch_HP_ON_OFF;
         R     "DB614_MH_State".MH_Status[2].Switch_HP_ON_OFF;
         R     "DB614_MH_State".MH_Status[3].Switch_HP_ON_OFF;
         R     "DB614_MH_State".MH_Status[4].Switch_HP_ON_OFF;
         R     "DB614_MH_State".MH_Status[5].Switch_HP_ON_OFF;
         R     "DB614_MH_State".MH_Status[6].Switch_HP_ON_OFF;
         R     "DB614_MH_State".MH_Status[7].Switch_HP_ON_OFF;
         R     "DB614_MH_State".MH_Status[8].Switch_HP_ON_OFF;
         R     "DB614_MH_State".MH_Status[9].Switch_HP_ON_OFF;
         R     "DB614_MH_State".MH_Status[10].Switch_HP_ON_OFF;
         R     "DB614_MH_State".MH_Status[11].Switch_HP_ON_OFF;
         R     "DB614_MH_State".MH_Status[12].Switch_HP_ON_OFF;
END_REGION

REGION Network 10: Shot preparation to start foaming cycle
   //For Interface 01:
   //
   //      O     "K_Vorbereitung_FT1"
   //      L     "DB761_Cylinder_Manager".CylinderMan_Ma[1].Preparation_Cylinder
   //      SI    "TM_Vorbereitung_SS01"
   //__________________________________________________________________
   //
   //    O     "TM_Vorbereitung_SS01"
   //    O     "TM_Vorbereitung_SS02"
   //    U     "DB619_State_MPart".Operationmode_Ma[1].Auto
         CLR;
         =     #Temp_ShotPreperation;
END_REGION

REGION Network 11: Detecting recirculation modes
         CALL  "FC012_Circulation"
         ( IN_OperationMode_Manual  := "DB619_State_MPart".Operationmode[1].Manual,
           IN_OperationMode_Auto    := "DB619_State_MPart".Operationmode[1].Auto,
           IN_OperationMode_active  := "DB619_State_MPart".Operationmode[1].Active,
           IN_Hydraulic_Switched_ON := "DB611_Hydraulic_State".MH_Hydraulic[1].Switch_Hydraulic_ON_OFF,
           IN_Hydraulic_OK          := "DB619_State_MPart".Machine[1].HydStartUp_finished,
           IN_LampTest              := "DB619_State_MPart".Operationmode[1].Lamptest,
           IN_Cycle_running         := "DB619_State_MPart".Cycle[1].running,
           IN_ShotPreparation_KK    := #Temp_ShotPreperation,
           IN_Fault_Level_1         := "DB009_Faults".Fault_State_Grp_1_M1,
           IN_Release_HP_Circ       := #Temp_Release_HP,
           IN_KK_in_PausingPos      := TRUE,  //"DB761_Cylinder_Manager".CylinderMan_Ma[1].Stop_to_Pause
           IN_Circulation_Timer     := "TM_Kreislauf_M1",
           IN_Runtime_Manual        := "DB700_Machine".Machine[1].Int_Runtime_Manual,
           IN_Breaktime_Manual      := "DB700_Machine".Machine[1].Int_Pausetime_Manual,
           IN_Runtime_Auto          := "DB700_Machine".Machine[1].Int_Runtime_Auto,
           IN_Breaktime_Auto        := "DB700_Machine".Machine[1].Int_Pausetime_Auto,
           IN_SWU_Release           := "DB619_State_MPart".SWU[1].SWU_released,
           OU_MesIntervallTimeNOK   := "DB820_Error_general".Machine[1].TimeValueIntervallNOK,
           IO_Status                := "DB619_State_MPart".Recirculation[1]
         );
   //
END_REGION

REGION Network 12: Activate indication high pressure cycle active
         L     0;
         T     "DB614_MH_State".MH_Status[1].State_HP;
         T     "DB614_MH_State".MH_Status[2].State_HP;
         T     "DB614_MH_State".MH_Status[3].State_HP;
         T     "DB614_MH_State".MH_Status[4].State_HP;
         T     "DB614_MH_State".MH_Status[5].State_HP;
         T     "DB614_MH_State".MH_Status[6].State_HP;
         T     "DB614_MH_State".MH_Status[7].State_HP;
         T     "DB614_MH_State".MH_Status[8].State_HP;
         T     "DB614_MH_State".MH_Status[9].State_HP;
         T     "DB614_MH_State".MH_Status[10].State_HP;
         T     "DB614_MH_State".MH_Status[11].State_HP;
         T     "DB614_MH_State".MH_Status[12].State_HP;

